   "Carrier_23_ActualSpeed" AT %IW1520 : Word;   // ACTUAL SPEED
   "Carrier_23_CarrierDriveAlarm" AT %IW1522 : Word;   // CARRIER DRIVE ALARM
   "Carrier_23_CarrierDriveWarning" AT %IW1524 : Word;   // CARRIER DRIVE WARNING
   "Carrier_24_Status" AT %IW1550 : Word;   // CARRIER STATUS WORD
   "Carrier_24_Status.0" AT %I1550.0 : Bool;   // HEARTBEAT
   "Carrier_24_Status.1" AT %I1550.1 : Bool;   // MANUAL
   "Carrier_24_Status.2" AT %I1550.2 : Bool;   // IN_AUTO
   "Carrier_24_Status.3" AT %I1550.3 : Bool;   // POSITIONING_COMPLETE
   "Carrier_24_Status.4" AT %I1550.4 : Bool;   // PRODUCTION HOLD
   "Carrier_24_Status.5" AT %I1550.5 : Bool;   // CARRIER MOVING FORWARD
   "Carrier_24_Status.6" AT %I1550.6 : Bool;   // CARRIER MOVING REVERSE
   "Carrier_24_Status.7" AT %I1550.7 : Bool;   // CARRIER FAULT
   "Carrier_24_Status.8" AT %I1551.0 : Bool;   // CRASH DETECT TRIPPED
   "Carrier_24_Status.9" AT %I1551.1 : Bool;
   "Carrier_24_Status.10" AT %I1551.2 : Bool;
   "Carrier_24_Status.11" AT %I1551.3 : Bool;
   "Carrier_24_Status.12" AT %I1551.4 : Bool;
   "Carrier_24_Status.13" AT %I1551.5 : Bool;
   "Carrier_24_Status.14" AT %I1551.6 : Bool;
   "Carrier_24_Status.15" AT %I1551.7 : Bool;
   "Carrier_24_SDCFaultCode" AT %IW1552 : Word;   // SDC FAULT CODE
   "Carrier_24_CarrierPosition" AT %ID1554 : DWord;   // CARRIER POSITION
   "Carrier_24_CarrierNumber" AT %IW1558 : Word;   // CARRIER NUMBER
   "Carrier_24_G120DControlWord" AT %IW1560 : Word;   // G120D_STW1_CONTROL
   "Carrier_24_G120DControlWord.0" AT %I1560.0 : Bool;   // Bit_00_ON
   "Carrier_24_G120DControlWord.1" AT %I1560.1 : Bool;   // Bit_01_AUS2_INH
   "Carrier_24_G120DControlWord.2" AT %I1560.2 : Bool;   // Bit_02_AUS3_STOP
   "Carrier_24_G120DControlWord.3" AT %I1560.3 : Bool;   // Bit_03_EN
   "Carrier_24_G120DControlWord.4" AT %I1560.4 : Bool;   // Bit_04_EN_RAMP
   "Carrier_24_G120DControlWord.5" AT %I1560.5 : Bool;   // Bit_05_START_RAMP
   "Carrier_24_G120DControlWord.6" AT %I1560.6 : Bool;   // Bit_06_SETPOINT
   "Carrier_24_G120DControlWord.7" AT %I1560.7 : Bool;   // Bit_07_RESET
   "Carrier_24_G120DControlWord.8" AT %I1561.0 : Bool;   // Bit_08_JOG_R
   "Carrier_24_G120DControlWord.9" AT %I1561.1 : Bool;   // Bit_09_JOG_L
   "Carrier_24_G120DControlWord.10" AT %I1561.2 : Bool;   // Bit_10_CONTR_PLC
   "Carrier_24_G120DControlWord.11" AT %I1561.3 : Bool;   // Bit_11_REVERSE
   "Carrier_24_G120DControlWord.12" AT %I1561.4 : Bool;   // Bit_12_BRAKE_RELEASE
   "Carrier_24_G120DControlWord.13" AT %I1561.5 : Bool;   // Bit_13_DDS
   "Carrier_24_G120DControlWord.14" AT %I1561.6 : Bool;   // Bit_14_DO0
   "Carrier_24_G120DControlWord.15" AT %I1561.7 : Bool;   // Bit_15_DO1
   "Carrier_24_G120DStatusWord" AT %IW1562 : Word;   // G120D_ZSW1_STATUS
   "Carrier_24_G120DStatusWord.0" AT %I1562.0 : Bool;   // Bit_00_READY_RUN
   "Carrier_24_G120DStatusWord.1" AT %I1562.1 : Bool;   // Bit_01_READY_ON
   "Carrier_24_G120DStatusWord.2" AT %I1562.2 : Bool;   // Bit_02_ENABLE
   "Carrier_24_G120DStatusWord.3" AT %I1562.3 : Bool;   // Bit_03_FAULT
   "Carrier_24_G120DStatusWord.4" AT %I1562.4 : Bool;   // Bit_04_OFF2
   "Carrier_24_G120DStatusWord.5" AT %I1562.5 : Bool;   // Bit_05_OFF3
   "Carrier_24_G120DStatusWord.6" AT %I1562.6 : Bool;   // Bit_06_LOCK_OUT
   "Carrier_24_G120DStatusWord.7" AT %I1562.7 : Bool;   // Bit_07_WARN
   "Carrier_24_G120DStatusWord.8" AT %I1563.0 : Bool;   // Bit_08_NO_DEVIATION
   "Carrier_24_G120DStatusWord.9" AT %I1563.1 : Bool;   // Bit_09_CONTR_PLC
   "Carrier_24_G120DStatusWord.10" AT %I1563.2 : Bool;   // Bit_10_F_MAX
   "Carrier_24_G120DStatusWord.11" AT %I1563.3 : Bool;   // Bit_11_LIMIT_REACHED
   "Carrier_24_G120DStatusWord.12" AT %I1563.4 : Bool;   // Bit_12_BRAKE_OPEN
   "Carrier_24_G120DStatusWord.13" AT %I1563.5 : Bool;   // Bit_13_NO_OVERTEMP
   "Carrier_24_G120DStatusWord.14" AT %I1563.6 : Bool;   // Bit_14_CW_CCW
   "Carrier_24_G120DStatusWord.15" AT %I1563.7 : Bool;   // Bit_15_OVERL
   "Carrier_24_Slot2_Input" AT %IW1564 : Word;   // SLOT 2 INPUT WORD
   "Carrier_24_CrashDetectSW" AT %I1564.0 : Bool;   // CRASH DETECT SW
   "Carrier_24_SpareSafetyInput(2_1)" AT %I1564.1 : Bool;   // SPARE SAFETY INPUT
   "Carrier_24_SpareSafetyInput(2_2)" AT %I1564.2 : Bool;   // SPARE SAFETY INPUT
   "Carrier_24_SpareSafetyInput(2_3)" AT %I1564.3 : Bool;   // SPARE SAFETY INPUT
   "Carrier_24_SpareSafetyInput(2_4)" AT %I1564.4 : Bool;   // SPARE SAFETY INPUT
   "Carrier_24_SpareSafetyInput(2_5)" AT %I1564.5 : Bool;   // SPARE SAFETY INPUT
   "Carrier_24_SpareSafetyInput(2_6)" AT %I1564.6 : Bool;   // SPARE SAFETY INPUT
   "Carrier_24_SpareSafetyInput(2_7)" AT %I1564.7 : Bool;   // SPARE SAFETY INPUT
   "Carrier_24_Slot3_SafetyOutput" AT %IW1565 : Word;   // SLOT 3 SAFETY OUTPUT WORD
   "Carrier_24_Crash_Detect_OK" AT %I1565.0 : Bool;   // CARRIER CRASH DETECT
   "Carrier_24_SpareSafetyOutput(3_1)" AT %I1565.1 : Bool;   // SPARE SAFETY OUTPUT
   "Carrier_24_SpareSafetyOutput(3_2)" AT %I1565.2 : Bool;   // SPARE SAFETY OUTPUT
   "Carrier_24_SpareSafetyOutput(3_3)" AT %I1565.3 : Bool;   // SPARE SAFETY OUTPUT
   "Carrier_24_SpareSafetyOutput(3_4)" AT %I1565.4 : Bool;   // SPARE SAFETY OUTPUT
   "Carrier_24_SpareSafetyOutput(3_5)" AT %I1565.5 : Bool;   // SPARE SAFETY OUTPUT
   "Carrier_24_SpareSafetyOutput(3_6)" AT %I1565.6 : Bool;   // SPARE SAFETY OUTPUT
   "Carrier_24_SpareSafetyOutput(3_7)" AT %I1565.7 : Bool;   // SPARE SAFETY OUTPUT
   "Carrier_24_Slot4_Input" AT %IW1566 : Word;   // SLOT 4 INPUT WORD
   "Carrier_24_480VPowerOn_MDCB1" AT %I1566.0 : Bool;   // 480 VAC POWER ON MDCB 1
   "Carrier_24_SpareInput(4_1)" AT %I1566.1 : Bool;   // SPARE INPUT
   "Carrier_24_SpareInput(4_2)" AT %I1566.2 : Bool;   // SPARE INPUT
   "Carrier_24_SitopSelectStatus" AT %I1566.3 : Bool;   // SITOP SELECT STATUS
   "Carrier_24_DCsupplyOnPSCB2" AT %I1566.4 : Bool;   // DC SUPPLY ON PSCB 2
   "Carrier_24_SpareInput(4_5)" AT %I1566.5 : Bool;   // SPARE INPUT
   "Carrier_24_SpareInput(4_6)" AT %I1566.6 : Bool;   // SPARE INPUT
   "Carrier_24_SpareInput(4_7)" AT %I1566.7 : Bool;   // SPARE INPUT
   "Carrier_24_PB1_ProdHoldLH" AT %I1567.0 : Bool;   // PB 1 PRODUCTION HOLD LH
   "Carrier_24_PB2_ResetLH" AT %I1567.1 : Bool;   // PB 2 RESET LH
   "Carrier_24_PB3_ProdHoldRH" AT %I1567.2 : Bool;   // PB 3 PRODUCTION HOLD RH
   "Carrier_24_PB4_ResetRH" AT %I1567.3 : Bool;   // PB 4 RESET RH
   "Carrier_24_SpareInput(4_14)" AT %I1567.4 : Bool;   // SPARE INPUT
   "Carrier_24_SpareInput(4_15)" AT %I1567.5 : Bool;   // SPARE INPUT
   "Carrier_24_SpareInput(4_16)" AT %I1567.6 : Bool;   // SPARE INPUT
   "Carrier_24_SpareInput(4_17)" AT %I1567.7 : Bool;   // SPARE INPUT
   "Carrier_24_Slot5_Output" AT %IW1568 : Word;   // SLOT 5 OUTPUT WORD
   "Carrier_24_IRD400_HMI_24VDC_ENABLE" AT %I1568.0 : Bool;   // IRD 400 PANEL HMI 24V DC POWER
   "Carrier_24_FaultLight_LH" AT %I1568.1 : Bool;   // FAULT LIGHT LH
   "Carrier_24_RunLight_LH" AT %I1568.2 : Bool;   // RUN LIGHT LH
   "Carrier_24_FaultLight_RH" AT %I1568.3 : Bool;   // FAULT LIGHT RH
   "Carrier_24_RunLight_RH" AT %I1568.4 : Bool;   // RUN LIGHT RH
   "Carrier_24_SpareOutput(5_5)" AT %I1568.5 : Bool;   // SPARE OUTPUT
   "Carrier_24_SpareOutput(5_6)" AT %I1568.6 : Bool;   // SPARE OUTPUT
   "Carrier_24_SpareOutput(5_7)" AT %I1568.7 : Bool;   // SPARE OUTPUT
   "Carrier_24_ActualSpeed" AT %IW1570 : Word;   // ACTUAL SPEED
   "Carrier_24_CarrierDriveAlarm" AT %IW1572 : Word;   // CARRIER DRIVE ALARM
   "Carrier_24_CarrierDriveWarning" AT %IW1574 : Word;   // CARRIER DRIVE WARNING
   "Carrier_25_Status" AT %IW1600 : Word;   // CARRIER STATUS WORD
   "Carrier_25_Status.0" AT %I1600.0 : Bool;   // HEARTBEAT
   "Carrier_25_Status.1" AT %I1600.1 : Bool;   // MANUAL
   "Carrier_25_Status.2" AT %I1600.2 : Bool;   // IN_AUTO
   "Carrier_25_Status.3" AT %I1600.3 : Bool;   // POSITIONING_COMPLETE
   "Carrier_25_Status.4" AT %I1600.4 : Bool;   // PRODUCTION HOLD
   "Carrier_25_Status.5" AT %I1600.5 : Bool;   // CARRIER MOVING FORWARD
   "Carrier_25_Status.6" AT %I1600.6 : Bool;   // CARRIER MOVING REVERSE
   "Carrier_25_Status.7" AT %I1600.7 : Bool;   // CARRIER FAULT
   "Carrier_25_Status.8" AT %I1601.0 : Bool;   // CRASH DETECT TRIPPED
   "Carrier_25_Status.9" AT %I1601.1 : Bool;
   "Carrier_25_Status.10" AT %I1601.2 : Bool;
   "Carrier_25_Status.11" AT %I1601.3 : Bool;
   "Carrier_25_Status.12" AT %I1601.4 : Bool;
   "Carrier_25_Status.13" AT %I1601.5 : Bool;
   "Carrier_25_Status.14" AT %I1601.6 : Bool;
   "Carrier_25_Status.15" AT %I1601.7 : Bool;
   "Carrier_25_SDCFaultCode" AT %IW1602 : Word;   // SDC FAULT CODE
   "Carrier_25_CarrierPosition" AT %ID1604 : DWord;   // CARRIER POSITION
   "Carrier_25_CarrierNumber" AT %IW1608 : Word;   // CARRIER NUMBER
   "Carrier_25_G120DControlWord" AT %IW1610 : Word;   // G120D_STW1_CONTROL
   "Carrier_25_G120DControlWord.0" AT %I1610.0 : Bool;   // Bit_00_ON
   "Carrier_25_G120DControlWord.1" AT %I1610.1 : Bool;   // Bit_01_AUS2_INH
   "Carrier_25_G120DControlWord.2" AT %I1610.2 : Bool;   // Bit_02_AUS3_STOP
   "Carrier_25_G120DControlWord.3" AT %I1610.3 : Bool;   // Bit_03_EN
   "Carrier_25_G120DControlWord.4" AT %I1610.4 : Bool;   // Bit_04_EN_RAMP
   "Carrier_25_G120DControlWord.5" AT %I1610.5 : Bool;   // Bit_05_START_RAMP
   "Carrier_25_G120DControlWord.6" AT %I1610.6 : Bool;   // Bit_06_SETPOINT
   "Carrier_25_G120DControlWord.7" AT %I1610.7 : Bool;   // Bit_07_RESET
   "Carrier_25_G120DControlWord.8" AT %I1611.0 : Bool;   // Bit_08_JOG_R
   "Carrier_25_G120DControlWord.9" AT %I1611.1 : Bool;   // Bit_09_JOG_L
   "Carrier_25_G120DControlWord.10" AT %I1611.2 : Bool;   // Bit_10_CONTR_PLC
   "Carrier_25_G120DControlWord.11" AT %I1611.3 : Bool;   // Bit_11_REVERSE
   "Carrier_25_G120DControlWord.12" AT %I1611.4 : Bool;   // Bit_12_BRAKE_RELEASE
   "Carrier_25_G120DControlWord.13" AT %I1611.5 : Bool;   // Bit_13_DDS
   "Carrier_25_G120DControlWord.14" AT %I1611.6 : Bool;   // Bit_14_DO0
   "Carrier_25_G120DControlWord.15" AT %I1611.7 : Bool;   // Bit_15_DO1
   "Carrier_25_G120DStatusWord" AT %IW1612 : Word;   // G120D_ZSW1_STATUS
   "Carrier_25_G120DStatusWord.0" AT %I1612.0 : Bool;   // Bit_00_READY_RUN
   "Carrier_25_G120DStatusWord.1" AT %I1612.1 : Bool;   // Bit_01_READY_ON
   "Carrier_25_G120DStatusWord.2" AT %I1612.2 : Bool;   // Bit_02_ENABLE
   "Carrier_25_G120DStatusWord.3" AT %I1612.3 : Bool;   // Bit_03_FAULT
   "Carrier_25_G120DStatusWord.4" AT %I1612.4 : Bool;   // Bit_04_OFF2
   "Carrier_25_G120DStatusWord.5" AT %I1612.5 : Bool;   // Bit_05_OFF3
   "Carrier_25_G120DStatusWord.6" AT %I1612.6 : Bool;   // Bit_06_LOCK_OUT
   "Carrier_25_G120DStatusWord.7" AT %I1612.7 : Bool;   // Bit_07_WARN
   "Carrier_25_G120DStatusWord.8" AT %I1613.0 : Bool;   // Bit_08_NO_DEVIATION
   "Carrier_25_G120DStatusWord.9" AT %I1613.1 : Bool;   // Bit_09_CONTR_PLC
   "Carrier_25_G120DStatusWord.10" AT %I1613.2 : Bool;   // Bit_10_F_MAX
   "Carrier_25_G120DStatusWord.11" AT %I1613.3 : Bool;   // Bit_11_LIMIT_REACHED
   "Carrier_25_G120DStatusWord.12" AT %I1613.4 : Bool;   // Bit_12_BRAKE_OPEN
   "Carrier_25_G120DStatusWord.13" AT %I1613.5 : Bool;   // Bit_13_NO_OVERTEMP
   "Carrier_25_G120DStatusWord.14" AT %I1613.6 : Bool;   // Bit_14_CW_CCW
   "Carrier_25_G120DStatusWord.15" AT %I1613.7 : Bool;   // Bit_15_OVERL
   "Carrier_25_Slot2_Input" AT %IW1614 : Word;   // SLOT 2 INPUT WORD
   "Carrier_25_CrashDetectSW" AT %I1614.0 : Bool;   // CRASH DETECT SW
   "Carrier_25_SpareSafetyInput(2_1)" AT %I1614.1 : Bool;   // SPARE SAFETY INPUT
   "Carrier_25_SpareSafetyInput(2_2)" AT %I1614.2 : Bool;   // SPARE SAFETY INPUT
   "Carrier_25_SpareSafetyInput(2_3)" AT %I1614.3 : Bool;   // SPARE SAFETY INPUT
   "Carrier_25_SpareSafetyInput(2_4)" AT %I1614.4 : Bool;   // SPARE SAFETY INPUT
   "Carrier_25_SpareSafetyInput(2_5)" AT %I1614.5 : Bool;   // SPARE SAFETY INPUT
   "Carrier_25_SpareSafetyInput(2_6)" AT %I1614.6 : Bool;   // SPARE SAFETY INPUT
   "Carrier_25_SpareSafetyInput(2_7)" AT %I1614.7 : Bool;   // SPARE SAFETY INPUT
   "Carrier_25_Slot3_SafetyOutput" AT %IW1615 : Word;   // SLOT 3 SAFETY OUTPUT WORD
   "Carrier_25_Crash_Detect_OK" AT %I1615.0 : Bool;   // CARRIER CRASH DETECT
   "Carrier_25_SpareSafetyOutput(3_1)" AT %I1615.1 : Bool;   // SPARE SAFETY OUTPUT
   "Carrier_25_SpareSafetyOutput(3_2)" AT %I1615.2 : Bool;   // SPARE SAFETY OUTPUT
   "Carrier_25_SpareSafetyOutput(3_3)" AT %I1615.3 : Bool;   // SPARE SAFETY OUTPUT
   "Carrier_25_SpareSafetyOutput(3_4)" AT %I1615.4 : Bool;   // SPARE SAFETY OUTPUT
   "Carrier_25_SpareSafetyOutput(3_5)" AT %I1615.5 : Bool;   // SPARE SAFETY OUTPUT
   "Carrier_25_SpareSafetyOutput(3_6)" AT %I1615.6 : Bool;   // SPARE SAFETY OUTPUT
   "Carrier_25_SpareSafetyOutput(3_7)" AT %I1615.7 : Bool;   // SPARE SAFETY OUTPUT
   "Carrier_25_Slot4_Input" AT %IW1616 : Word;   // SLOT 4 INPUT WORD
   "Carrier_25_480VPowerOn_MDCB1" AT %I1616.0 : Bool;   // 480 VAC POWER ON MDCB 1
   "Carrier_25_SpareInput(4_1)" AT %I1616.1 : Bool;   // SPARE INPUT
   "Carrier_25_SpareInput(4_2)" AT %I1616.2 : Bool;   // SPARE INPUT
   "Carrier_25_SitopSelectStatus" AT %I1616.3 : Bool;   // SITOP SELECT STATUS
   "Carrier_25_DCsupplyOnPSCB2" AT %I1616.4 : Bool;   // DC SUPPLY ON PSCB 2
   "Carrier_25_SpareInput(4_5)" AT %I1616.5 : Bool;   // SPARE INPUT
   "Carrier_25_SpareInput(4_6)" AT %I1616.6 : Bool;   // SPARE INPUT
   "Carrier_25_SpareInput(4_7)" AT %I1616.7 : Bool;   // SPARE INPUT
   "Carrier_25_PB1_ProdHoldLH" AT %I1617.0 : Bool;   // PB 1 PRODUCTION HOLD LH
   "Carrier_25_PB2_ResetLH" AT %I1617.1 : Bool;   // PB 2 RESET LH
   "Carrier_25_PB3_ProdHoldRH" AT %I1617.2 : Bool;   // PB 3 PRODUCTION HOLD RH
   "Carrier_25_PB4_ResetRH" AT %I1617.3 : Bool;   // PB 4 RESET RH
   "Carrier_25_SpareInput(4_14)" AT %I1617.4 : Bool;   // SPARE INPUT
   "Carrier_25_SpareInput(4_15)" AT %I1617.5 : Bool;   // SPARE INPUT
   "Carrier_25_SpareInput(4_16)" AT %I1617.6 : Bool;   // SPARE INPUT
   "Carrier_25_SpareInput(4_17)" AT %I1617.7 : Bool;   // SPARE INPUT
   "Carrier_25_Slot5_Output" AT %IW1618 : Word;   // SLOT 5 OUTPUT WORD
   "Carrier_25_IRD400_HMI_24VDC_ENABLE" AT %I1618.0 : Bool;   // IRD 400 PANEL HMI 24V DC POWER
   "Carrier_25_FaultLight_LH" AT %I1618.1 : Bool;   // FAULT LIGHT LH
   "Carrier_25_RunLight_LH" AT %I1618.2 : Bool;   // RUN LIGHT LH
   "Carrier_25_FaultLight_RH" AT %I1618.3 : Bool;   // FAULT LIGHT RH
   "Carrier_25_RunLight_RH" AT %I1618.4 : Bool;   // RUN LIGHT RH
   "Carrier_25_SpareOutput(5_5)" AT %I1618.5 : Bool;   // SPARE OUTPUT
   "Carrier_25_SpareOutput(5_6)" AT %I1618.6 : Bool;   // SPARE OUTPUT
   "Carrier_25_SpareOutput(5_7)" AT %I1618.7 : Bool;   // SPARE OUTPUT
   "Carrier_25_ActualSpeed" AT %IW1620 : Word;   // ACTUAL SPEED
   "Carrier_25_CarrierDriveAlarm" AT %IW1622 : Word;   // CARRIER DRIVE ALARM
   "Carrier_25_CarrierDriveWarning" AT %IW1624 : Word;   // CARRIER DRIVE WARNING
   "Carrier_26_Status" AT %IW1650 : Word;   // CARRIER STATUS WORD
   "Carrier_26_Status.0" AT %I1650.0 : Bool;   // HEARTBEAT
   "Carrier_26_Status.1" AT %I1650.1 : Bool;   // MANUAL
   "Carrier_26_Status.2" AT %I1650.2 : Bool;   // IN_AUTO
   "Carrier_26_Status.3" AT %I1650.3 : Bool;   // POSITIONING_COMPLETE
   "Carrier_26_Status.4" AT %I1650.4 : Bool;   // PRODUCTION HOLD
   "Carrier_26_Status.5" AT %I1650.5 : Bool;   // CARRIER MOVING FORWARD
   "Carrier_26_Status.6" AT %I1650.6 : Bool;   // CARRIER MOVING REVERSE
   "Carrier_26_Status.7" AT %I1650.7 : Bool;   // CARRIER FAULT
   "Carrier_26_Status.8" AT %I1651.0 : Bool;   // CRASH DETECT TRIPPED
   "Carrier_26_Status.9" AT %I1651.1 : Bool;
   "Carrier_26_Status.10" AT %I1651.2 : Bool;
   "Carrier_26_Status.11" AT %I1651.3 : Bool;
   "Carrier_26_Status.12" AT %I1651.4 : Bool;
   "Carrier_26_Status.13" AT %I1651.5 : Bool;
   "Carrier_26_Status.14" AT %I1651.6 : Bool;
   "Carrier_26_Status.15" AT %I1651.7 : Bool;
   "Carrier_26_SDCFaultCode" AT %IW1652 : Word;   // SDC FAULT CODE
   "Carrier_26_CarrierPosition" AT %ID1654 : DWord;   // CARRIER POSITION
   "Carrier_26_CarrierNumber" AT %IW1658 : Word;   // CARRIER NUMBER
   "Carrier_26_G120DControlWord" AT %IW1660 : Word;   // G120D_STW1_CONTROL
   "Carrier_26_G120DControlWord.0" AT %I1660.0 : Bool;   // Bit_00_ON
   "Carrier_26_G120DControlWord.1" AT %I1660.1 : Bool;   // Bit_01_AUS2_INH
   "Carrier_26_G120DControlWord.2" AT %I1660.2 : Bool;   // Bit_02_AUS3_STOP
   "Carrier_26_G120DControlWord.3" AT %I1660.3 : Bool;   // Bit_03_EN
   "Carrier_26_G120DControlWord.4" AT %I1660.4 : Bool;   // Bit_04_EN_RAMP
   "Carrier_26_G120DControlWord.5" AT %I1660.5 : Bool;   // Bit_05_START_RAMP
   "Carrier_26_G120DControlWord.6" AT %I1660.6 : Bool;   // Bit_06_SETPOINT
   "Carrier_26_G120DControlWord.7" AT %I1660.7 : Bool;   // Bit_07_RESET
   "Carrier_26_G120DControlWord.8" AT %I1661.0 : Bool;   // Bit_08_JOG_R
   "Carrier_26_G120DControlWord.9" AT %I1661.1 : Bool;   // Bit_09_JOG_L
   "Carrier_26_G120DControlWord.10" AT %I1661.2 : Bool;   // Bit_10_CONTR_PLC
   "Carrier_26_G120DControlWord.11" AT %I1661.3 : Bool;   // Bit_11_REVERSE
   "Carrier_26_G120DControlWord.12" AT %I1661.4 : Bool;   // Bit_12_BRAKE_RELEASE
   "Carrier_26_G120DControlWord.13" AT %I1661.5 : Bool;   // Bit_13_DDS
   "Carrier_26_G120DControlWord.14" AT %I1661.6 : Bool;   // Bit_14_DO0
   "Carrier_26_G120DControlWord.15" AT %I1661.7 : Bool;   // Bit_15_DO1
   "Carrier_26_G120DStatusWord" AT %IW1662 : Word;   // G120D_ZSW1_STATUS
   "Carrier_26_G120DStatusWord.0" AT %I1662.0 : Bool;   // Bit_00_READY_RUN
   "Carrier_26_G120DStatusWord.1" AT %I1662.1 : Bool;   // Bit_01_READY_ON
   "Carrier_26_G120DStatusWord.2" AT %I1662.2 : Bool;   // Bit_02_ENABLE
   "Carrier_26_G120DStatusWord.3" AT %I1662.3 : Bool;   // Bit_03_FAULT
   "Carrier_26_G120DStatusWord.4" AT %I1662.4 : Bool;   // Bit_04_OFF2
   "Carrier_26_G120DStatusWord.5" AT %I1662.5 : Bool;   // Bit_05_OFF3
   "Carrier_26_G120DStatusWord.6" AT %I1662.6 : Bool;   // Bit_06_LOCK_OUT
   "Carrier_26_G120DStatusWord.7" AT %I1662.7 : Bool;   // Bit_07_WARN
   "Carrier_26_G120DStatusWord.8" AT %I1663.0 : Bool;   // Bit_08_NO_DEVIATION
   "Carrier_26_G120DStatusWord.9" AT %I1663.1 : Bool;   // Bit_09_CONTR_PLC
   "Carrier_26_G120DStatusWord.10" AT %I1663.2 : Bool;   // Bit_10_F_MAX
   "Carrier_26_G120DStatusWord.11" AT %I1663.3 : Bool;   // Bit_11_LIMIT_REACHED
   "Carrier_26_G120DStatusWord.12" AT %I1663.4 : Bool;   // Bit_12_BRAKE_OPEN
   "Carrier_26_G120DStatusWord.13" AT %I1663.5 : Bool;   // Bit_13_NO_OVERTEMP
   "Carrier_26_G120DStatusWord.14" AT %I1663.6 : Bool;   // Bit_14_CW_CCW
   "Carrier_26_G120DStatusWord.15" AT %I1663.7 : Bool;   // Bit_15_OVERL
   "Carrier_26_Slot2_Input" AT %IW1664 : Word;   // SLOT 2 INPUT WORD
   "Carrier_26_CrashDetectSW" AT %I1664.0 : Bool;   // CRASH DETECT SW
   "Carrier_26_SpareSafetyInput(2_1)" AT %I1664.1 : Bool;   // SPARE SAFETY INPUT
   "Carrier_26_SpareSafetyInput(2_2)" AT %I1664.2 : Bool;   // SPARE SAFETY INPUT
   "Carrier_26_SpareSafetyInput(2_3)" AT %I1664.3 : Bool;   // SPARE SAFETY INPUT
   "Carrier_26_SpareSafetyInput(2_4)" AT %I1664.4 : Bool;   // SPARE SAFETY INPUT
   "Carrier_26_SpareSafetyInput(2_5)" AT %I1664.5 : Bool;   // SPARE SAFETY INPUT
   "Carrier_26_SpareSafetyInput(2_6)" AT %I1664.6 : Bool;   // SPARE SAFETY INPUT
   "Carrier_26_SpareSafetyInput(2_7)" AT %I1664.7 : Bool;   // SPARE SAFETY INPUT
   "Carrier_26_Slot3_SafetyOutput" AT %IW1665 : Word;   // SLOT 3 SAFETY OUTPUT WORD
   "Carrier_26_Crash_Detect_OK" AT %I1665.0 : Bool;   // CARRIER CRASH DETECT
   "Carrier_26_SpareSafetyOutput(3_1)" AT %I1665.1 : Bool;   // SPARE SAFETY OUTPUT
   "Carrier_26_SpareSafetyOutput(3_2)" AT %I1665.2 : Bool;   // SPARE SAFETY OUTPUT
   "Carrier_26_SpareSafetyOutput(3_3)" AT %I1665.3 : Bool;   // SPARE SAFETY OUTPUT
   "Carrier_26_SpareSafetyOutput(3_4)" AT %I1665.4 : Bool;   // SPARE SAFETY OUTPUT
   "Carrier_26_SpareSafetyOutput(3_5)" AT %I1665.5 : Bool;   // SPARE SAFETY OUTPUT
   "Carrier_26_SpareSafetyOutput(3_6)" AT %I1665.6 : Bool;   // SPARE SAFETY OUTPUT
   "Carrier_26_SpareSafetyOutput(3_7)" AT %I1665.7 : Bool;   // SPARE SAFETY OUTPUT
   "Carrier_26_Slot4_Input" AT %IW1666 : Word;   // SLOT 4 INPUT WORD
   "Carrier_26_480VPowerOn_MDCB1" AT %I1666.0 : Bool;   // 480 VAC POWER ON MDCB 1
   "Carrier_26_SpareInput(4_1)" AT %I1666.1 : Bool;   // SPARE INPUT
   "Carrier_26_SpareInput(4_2)" AT %I1666.2 : Bool;   // SPARE INPUT
   "Carrier_26_SitopSelectStatus" AT %I1666.3 : Bool;   // SITOP SELECT STATUS
   "Carrier_26_DCsupplyOnPSCB2" AT %I1666.4 : Bool;   // DC SUPPLY ON PSCB 2
   "Carrier_26_SpareInput(4_5)" AT %I1666.5 : Bool;   // SPARE INPUT
   "Carrier_26_SpareInput(4_6)" AT %I1666.6 : Bool;   // SPARE INPUT
   "Carrier_26_SpareInput(4_7)" AT %I1666.7 : Bool;   // SPARE INPUT
   "Carrier_26_PB1_ProdHoldLH" AT %I1667.0 : Bool;   // PB 1 PRODUCTION HOLD LH
   "Carrier_26_PB2_ResetLH" AT %I1667.1 : Bool;   // PB 2 RESET LH
   "Carrier_26_PB3_ProdHoldRH" AT %I1667.2 : Bool;   // PB 3 PRODUCTION HOLD RH
   "Carrier_26_PB4_ResetRH" AT %I1667.3 : Bool;   // PB 4 RESET RH
   "Carrier_26_SpareInput(4_14)" AT %I1667.4 : Bool;   // SPARE INPUT
   "Carrier_26_SpareInput(4_15)" AT %I1667.5 : Bool;   // SPARE INPUT
   "Carrier_26_SpareInput(4_16)" AT %I1667.6 : Bool;   // SPARE INPUT
   "Carrier_26_SpareInput(4_17)" AT %I1667.7 : Bool;   // SPARE INPUT
   "Carrier_26_Slot5_Output" AT %IW1668 : Word;   // SLOT 5 OUTPUT WORD
   "Carrier_26_IRD400_HMI_24VDC_ENABLE" AT %I1668.0 : Bool;   // IRD 400 PANEL HMI 24V DC POWER
   "Carrier_26_FaultLight_LH" AT %I1668.1 : Bool;   // FAULT LIGHT LH
   "Carrier_26_RunLight_LH" AT %I1668.2 : Bool;   // RUN LIGHT LH
   "Carrier_26_FaultLight_RH" AT %I1668.3 : Bool;   // FAULT LIGHT RH
   "Carrier_26_RunLight_RH" AT %I1668.4 : Bool;   // RUN LIGHT RH
   "Carrier_26_SpareOutput(5_5)" AT %I1668.5 : Bool;   // SPARE OUTPUT
   "Carrier_26_SpareOutput(5_6)" AT %I1668.6 : Bool;   // SPARE OUTPUT
   "Carrier_26_SpareOutput(5_7)" AT %I1668.7 : Bool;   // SPARE OUTPUT
   "Carrier_26_ActualSpeed" AT %IW1670 : Word;   // ACTUAL SPEED
   "Carrier_26_CarrierDriveAlarm" AT %IW1672 : Word;   // CARRIER DRIVE ALARM
   "Carrier_26_CarrierDriveWarning" AT %IW1674 : Word;   // CARRIER DRIVE WARNING
   "Carrier_27_Status" AT %IW1700 : Word;   // CARRIER STATUS WORD
   "Carrier_27_Status.0" AT %I1700.0 : Bool;   // HEARTBEAT
   "Carrier_27_Status.1" AT %I1700.1 : Bool;   // MANUAL
   "Carrier_27_Status.2" AT %I1700.2 : Bool;   // IN_AUTO
   "Carrier_27_Status.3" AT %I1700.3 : Bool;   // POSITIONING_COMPLETE
   "Carrier_27_Status.4" AT %I1700.4 : Bool;   // PRODUCTION HOLD
   "Carrier_27_Status.5" AT %I1700.5 : Bool;   // CARRIER MOVING FORWARD
   "Carrier_27_Status.6" AT %I1700.6 : Bool;   // CARRIER MOVING REVERSE
   "Carrier_27_Status.7" AT %I1700.7 : Bool;   // CARRIER FAULT
   "Carrier_27_Status.8" AT %I1701.0 : Bool;   // CRASH DETECT TRIPPED
   "Carrier_27_Status.9" AT %I1701.1 : Bool;
   "Carrier_27_Status.10" AT %I1701.2 : Bool;
   "Carrier_27_Status.11" AT %I1701.3 : Bool;
   "Carrier_27_Status.12" AT %I1701.4 : Bool;
   "Carrier_27_Status.13" AT %I1701.5 : Bool;
   "Carrier_27_Status.14" AT %I1701.6 : Bool;
   "Carrier_27_Status.15" AT %I1701.7 : Bool;
   "Carrier_27_SDCFaultCode" AT %IW1702 : Word;   // SDC FAULT CODE
   "Carrier_27_CarrierPosition" AT %ID1704 : DWord;   // CARRIER POSITION
   "Carrier_27_CarrierNumber" AT %IW1708 : Word;   // CARRIER NUMBER
   "Carrier_27_G120DControlWord" AT %IW1710 : Word;   // G120D_STW1_CONTROL
   "Carrier_27_G120DControlWord.0" AT %I1710.0 : Bool;   // Bit_00_ON
   "Carrier_27_G120DControlWord.1" AT %I1710.1 : Bool;   // Bit_01_AUS2_INH
   "Carrier_27_G120DControlWord.2" AT %I1710.2 : Bool;   // Bit_02_AUS3_STOP
   "Carrier_27_G120DControlWord.3" AT %I1710.3 : Bool;   // Bit_03_EN
   "Carrier_27_G120DControlWord.4" AT %I1710.4 : Bool;   // Bit_04_EN_RAMP
   "Carrier_27_G120DControlWord.5" AT %I1710.5 : Bool;   // Bit_05_START_RAMP
   "Carrier_27_G120DControlWord.6" AT %I1710.6 : Bool;   // Bit_06_SETPOINT
   "Carrier_27_G120DControlWord.7" AT %I1710.7 : Bool;   // Bit_07_RESET
   "Carrier_27_G120DControlWord.8" AT %I1711.0 : Bool;   // Bit_08_JOG_R
   "Carrier_27_G120DControlWord.9" AT %I1711.1 : Bool;   // Bit_09_JOG_L
   "Carrier_27_G120DControlWord.10" AT %I1711.2 : Bool;   // Bit_10_CONTR_PLC
   "Carrier_27_G120DControlWord.11" AT %I1711.3 : Bool;   // Bit_11_REVERSE
   "Carrier_27_G120DControlWord.12" AT %I1711.4 : Bool;   // Bit_12_BRAKE_RELEASE
   "Carrier_27_G120DControlWord.13" AT %I1711.5 : Bool;   // Bit_13_DDS
   "Carrier_27_G120DControlWord.14" AT %I1711.6 : Bool;   // Bit_14_DO0
   "Carrier_27_G120DControlWord.15" AT %I1711.7 : Bool;   // Bit_15_DO1
   "Carrier_27_G120DStatusWord" AT %IW1712 : Word;   // G120D_ZSW1_STATUS
   "Carrier_27_G120DStatusWord.0" AT %I1712.0 : Bool;   // Bit_00_READY_RUN
   "Carrier_27_G120DStatusWord.1" AT %I1712.1 : Bool;   // Bit_01_READY_ON
   "Carrier_27_G120DStatusWord.2" AT %I1712.2 : Bool;   // Bit_02_ENABLE
   "Carrier_27_G120DStatusWord.3" AT %I1712.3 : Bool;   // Bit_03_FAULT
   "Carrier_27_G120DStatusWord.4" AT %I1712.4 : Bool;   // Bit_04_OFF2
   "Carrier_27_G120DStatusWord.5" AT %I1712.5 : Bool;   // Bit_05_OFF3
   "Carrier_27_G120DStatusWord.6" AT %I1712.6 : Bool;   // Bit_06_LOCK_OUT
   "Carrier_27_G120DStatusWord.7" AT %I1712.7 : Bool;   // Bit_07_WARN
   "Carrier_27_G120DStatusWord.8" AT %I1713.0 : Bool;   // Bit_08_NO_DEVIATION
   "Carrier_27_G120DStatusWord.9" AT %I1713.1 : Bool;   // Bit_09_CONTR_PLC
   "Carrier_27_G120DStatusWord.10" AT %I1713.2 : Bool;   // Bit_10_F_MAX
   "Carrier_27_G120DStatusWord.11" AT %I1713.3 : Bool;   // Bit_11_LIMIT_REACHED
   "Carrier_27_G120DStatusWord.12" AT %I1713.4 : Bool;   // Bit_12_BRAKE_OPEN
   "Carrier_27_G120DStatusWord.13" AT %I1713.5 : Bool;   // Bit_13_NO_OVERTEMP
   "Carrier_27_G120DStatusWord.14" AT %I1713.6 : Bool;   // Bit_14_CW_CCW
   "Carrier_27_G120DStatusWord.15" AT %I1713.7 : Bool;   // Bit_15_OVERL
   "Carrier_27_Slot2_Input" AT %IW1714 : Word;   // SLOT 2 INPUT WORD
   "Carrier_27_CrashDetectSW" AT %I1714.0 : Bool;   // CRASH DETECT SW
   "Carrier_27_SpareSafetyInput(2_1)" AT %I1714.1 : Bool;   // SPARE SAFETY INPUT
   "Carrier_27_SpareSafetyInput(2_2)" AT %I1714.2 : Bool;   // SPARE SAFETY INPUT
   "Carrier_27_SpareSafetyInput(2_3)" AT %I1714.3 : Bool;   // SPARE SAFETY INPUT
   "Carrier_27_SpareSafetyInput(2_4)" AT %I1714.4 : Bool;   // SPARE SAFETY INPUT
   "Carrier_27_SpareSafetyInput(2_5)" AT %I1714.5 : Bool;   // SPARE SAFETY INPUT
   "Carrier_27_SpareSafetyInput(2_6)" AT %I1714.6 : Bool;   // SPARE SAFETY INPUT
   "Carrier_27_SpareSafetyInput(2_7)" AT %I1714.7 : Bool;   // SPARE SAFETY INPUT
   "Carrier_27_Slot3_SafetyOutput" AT %IW1715 : Word;   // SLOT 3 SAFETY OUTPUT WORD
   "Carrier_27_Crash_Detect_OK" AT %I1715.0 : Bool;   // CARRIER CRASH DETECT
   "Carrier_27_SpareSafetyOutput(3_1)" AT %I1715.1 : Bool;   // SPARE SAFETY OUTPUT
   "Carrier_27_SpareSafetyOutput(3_2)" AT %I1715.2 : Bool;   // SPARE SAFETY OUTPUT
   "Carrier_27_SpareSafetyOutput(3_3)" AT %I1715.3 : Bool;   // SPARE SAFETY OUTPUT
   "Carrier_27_SpareSafetyOutput(3_4)" AT %I1715.4 : Bool;   // SPARE SAFETY OUTPUT
   "Carrier_27_SpareSafetyOutput(3_5)" AT %I1715.5 : Bool;   // SPARE SAFETY OUTPUT
   "Carrier_27_SpareSafetyOutput(3_6)" AT %I1715.6 : Bool;   // SPARE SAFETY OUTPUT
   "Carrier_27_SpareSafetyOutput(3_7)" AT %I1715.7 : Bool;   // SPARE SAFETY OUTPUT
   "Carrier_27_Slot4_Input" AT %IW1716 : Word;   // SLOT 4 INPUT WORD
   "Carrier_27_480VPowerOn_MDCB1" AT %I1716.0 : Bool;   // 480 VAC POWER ON MDCB 1
   "Carrier_27_SpareInput(4_1)" AT %I1716.1 : Bool;   // SPARE INPUT
   "Carrier_27_SpareInput(4_2)" AT %I1716.2 : Bool;   // SPARE INPUT
   "Carrier_27_SitopSelectStatus" AT %I1716.3 : Bool;   // SITOP SELECT STATUS
   "Carrier_27_DCsupplyOnPSCB2" AT %I1716.4 : Bool;   // DC SUPPLY ON PSCB 2
   "Carrier_27_SpareInput(4_5)" AT %I1716.5 : Bool;   // SPARE INPUT
   "Carrier_27_SpareInput(4_6)" AT %I1716.6 : Bool;   // SPARE INPUT
   "Carrier_27_SpareInput(4_7)" AT %I1716.7 : Bool;   // SPARE INPUT
   "Carrier_27_PB1_ProdHoldLH" AT %I1717.0 : Bool;   // PB 1 PRODUCTION HOLD LH
   "Carrier_27_PB2_ResetLH" AT %I1717.1 : Bool;   // PB 2 RESET LH
   "Carrier_27_PB3_ProdHoldRH" AT %I1717.2 : Bool;   // PB 3 PRODUCTION HOLD RH
   "Carrier_27_PB4_ResetRH" AT %I1717.3 : Bool;   // PB 4 RESET RH
   "Carrier_27_SpareInput(4_14)" AT %I1717.4 : Bool;   // SPARE INPUT
   "Carrier_27_SpareInput(4_15)" AT %I1717.5 : Bool;   // SPARE INPUT
   "Carrier_27_SpareInput(4_16)" AT %I1717.6 : Bool;   // SPARE INPUT
   "Carrier_27_SpareInput(4_17)" AT %I1717.7 : Bool;   // SPARE INPUT
   "Carrier_27_Slot5_Output" AT %IW1718 : Word;   // SLOT 5 OUTPUT WORD
   "Carrier_27_IRD400_HMI_24VDC_ENABLE" AT %I1718.0 : Bool;   // IRD 400 PANEL HMI 24V DC POWER
   "Carrier_27_FaultLight_LH" AT %I1718.1 : Bool;   // FAULT LIGHT LH
   "Carrier_27_RunLight_LH" AT %I1718.2 : Bool;   // RUN LIGHT LH
   "Carrier_27_FaultLight_RH" AT %I1718.3 : Bool;   // FAULT LIGHT RH
   "Carrier_27_RunLight_RH" AT %I1718.4 : Bool;   // RUN LIGHT RH
   "Carrier_27_SpareOutput(5_5)" AT %I1718.5 : Bool;   // SPARE OUTPUT
   "Carrier_27_SpareOutput(5_6)" AT %I1718.6 : Bool;   // SPARE OUTPUT
   "Carrier_27_SpareOutput(5_7)" AT %I1718.7 : Bool;   // SPARE OUTPUT
   "Carrier_27_ActualSpeed" AT %IW1720 : Word;   // ACTUAL SPEED
   "Carrier_27_CarrierDriveAlarm" AT %IW1722 : Word;   // CARRIER DRIVE ALARM
   "Carrier_27_CarrierDriveWarning" AT %IW1724 : Word;   // CARRIER DRIVE WARNING
   "Carrier_28_Status" AT %IW1750 : Word;   // CARRIER STATUS WORD
   "Carrier_28_Status.0" AT %I1750.0 : Bool;   // HEARTBEAT
   "Carrier_28_Status.1" AT %I1750.1 : Bool;   // MANUAL
   "Carrier_28_Status.2" AT %I1750.2 : Bool;   // IN_AUTO
   "Carrier_28_Status.3" AT %I1750.3 : Bool;   // POSITIONING_COMPLETE
   "Carrier_28_Status.4" AT %I1750.4 : Bool;   // PRODUCTION HOLD
   "Carrier_28_Status.5" AT %I1750.5 : Bool;   // CARRIER MOVING FORWARD
   "Carrier_28_Status.6" AT %I1750.6 : Bool;   // CARRIER MOVING REVERSE
   "Carrier_28_Status.7" AT %I1750.7 : Bool;   // CARRIER FAULT
   "Carrier_28_Status.8" AT %I1751.0 : Bool;   // CRASH DETECT TRIPPED
   "Carrier_28_Status.9" AT %I1751.1 : Bool;
   "Carrier_28_Status.10" AT %I1751.2 : Bool;
   "Carrier_28_Status.11" AT %I1751.3 : Bool;
   "Carrier_28_Status.12" AT %I1751.4 : Bool;
   "Carrier_28_Status.13" AT %I1751.5 : Bool;
   "Carrier_28_Status.14" AT %I1751.6 : Bool;
   "Carrier_28_Status.15" AT %I1751.7 : Bool;
   "Carrier_28_SDCFaultCode" AT %IW1752 : Word;   // SDC FAULT CODE
   "Carrier_28_CarrierPosition" AT %ID1754 : DWord;   // CARRIER POSITION
   "Carrier_28_CarrierNumber" AT %IW1758 : Word;   // CARRIER NUMBER
   "Carrier_28_G120DControlWord" AT %IW1760 : Word;   // G120D_STW1_CONTROL
   "Carrier_28_G120DControlWord.0" AT %I1760.0 : Bool;   // Bit_00_ON
   "Carrier_28_G120DControlWord.1" AT %I1760.1 : Bool;   // Bit_01_AUS2_INH
   "Carrier_28_G120DControlWord.2" AT %I1760.2 : Bool;   // Bit_02_AUS3_STOP
   "Carrier_28_G120DControlWord.3" AT %I1760.3 : Bool;   // Bit_03_EN
   "Carrier_28_G120DControlWord.4" AT %I1760.4 : Bool;   // Bit_04_EN_RAMP
   "Carrier_28_G120DControlWord.5" AT %I1760.5 : Bool;   // Bit_05_START_RAMP
   "Carrier_28_G120DControlWord.6" AT %I1760.6 : Bool;   // Bit_06_SETPOINT
   "Carrier_28_G120DControlWord.7" AT %I1760.7 : Bool;   // Bit_07_RESET
   "Carrier_28_G120DControlWord.8" AT %I1761.0 : Bool;   // Bit_08_JOG_R
   "Carrier_28_G120DControlWord.9" AT %I1761.1 : Bool;   // Bit_09_JOG_L
   "Carrier_28_G120DControlWord.10" AT %I1761.2 : Bool;   // Bit_10_CONTR_PLC
   "Carrier_28_G120DControlWord.11" AT %I1761.3 : Bool;   // Bit_11_REVERSE
   "Carrier_28_G120DControlWord.12" AT %I1761.4 : Bool;   // Bit_12_BRAKE_RELEASE
   "Carrier_28_G120DControlWord.13" AT %I1761.5 : Bool;   // Bit_13_DDS
   "Carrier_28_G120DControlWord.14" AT %I1761.6 : Bool;   // Bit_14_DO0
   "Carrier_28_G120DControlWord.15" AT %I1761.7 : Bool;   // Bit_15_DO1
   "Carrier_28_G120DStatusWord" AT %IW1762 : Word;   // G120D_ZSW1_STATUS
   "Carrier_28_G120DStatusWord.0" AT %I1762.0 : Bool;   // Bit_00_READY_RUN
   "Carrier_28_G120DStatusWord.1" AT %I1762.1 : Bool;   // Bit_01_READY_ON
   "Carrier_28_G120DStatusWord.2" AT %I1762.2 : Bool;   // Bit_02_ENABLE
   "Carrier_28_G120DStatusWord.3" AT %I1762.3 : Bool;   // Bit_03_FAULT
   "Carrier_28_G120DStatusWord.4" AT %I1762.4 : Bool;   // Bit_04_OFF2
   "Carrier_28_G120DStatusWord.5" AT %I1762.5 : Bool;   // Bit_05_OFF3
   "Carrier_28_G120DStatusWord.6" AT %I1762.6 : Bool;   // Bit_06_LOCK_OUT
   "Carrier_28_G120DStatusWord.7" AT %I1762.7 : Bool;   // Bit_07_WARN
   "Carrier_28_G120DStatusWord.8" AT %I1763.0 : Bool;   // Bit_08_NO_DEVIATION
   "Carrier_28_G120DStatusWord.9" AT %I1763.1 : Bool;   // Bit_09_CONTR_PLC
   "Carrier_28_G120DStatusWord.10" AT %I1763.2 : Bool;   // Bit_10_F_MAX
   "Carrier_28_G120DStatusWord.11" AT %I1763.3 : Bool;   // Bit_11_LIMIT_REACHED
   "Carrier_28_G120DStatusWord.12" AT %I1763.4 : Bool;   // Bit_12_BRAKE_OPEN
   "Carrier_28_G120DStatusWord.13" AT %I1763.5 : Bool;   // Bit_13_NO_OVERTEMP
   "Carrier_28_G120DStatusWord.14" AT %I1763.6 : Bool;   // Bit_14_CW_CCW
   "Carrier_28_G120DStatusWord.15" AT %I1763.7 : Bool;   // Bit_15_OVERL
   "Carrier_28_Slot2_Input" AT %IW1764 : Word;   // SLOT 2 INPUT WORD
   "Carrier_28_CrashDetectSW" AT %I1764.0 : Bool;   // CRASH DETECT SW
